         dHeadFireONDelay_cmm_H7 : DInt;   // Head#x fire ON delay [mm/100] {mm/100|mm|-50|50|O} / Head #7 fire ON delay [mm/100] {mm/100|mm|-50|50|O}
         dHeadFireOFFDelay_cmm_H7 : DInt;   // Head#x fire OFF delay [mm/100] {mm/100|mm|-50|50|O} / Head #7 fire OFF delay [mm/100] {mm/100|mm|-50|50|O}
         dHeadPressure_mN_H7 : DInt;   // Head#x pressure value [N/1000] {N/1000|N|16|180|O} / Head #7 pressure value [N/1000] {N/1000|N|16|180|O}
         dHeadFireONReaction_ms_H8 : DInt;   // Head#x fire ON reaction time [ms] {ms|s|0|1|M} / Head #8 fire ON reaction time [ms] {ms|s|0|1|M}
         dHeadFireOFFReaction_ms_H8 : DInt;   // Head#x fire OFF reaction time [ms] {ms|s|0|1|M} / Head #8 fire OFF reaction time [ms] {ms|s|0|1|M}
         dHeadOilONDelay_ms_H8 : DInt;   // Head#x Oil ON delay [ms]{ms|s|-2|2|O} / Head #8 Oil ON delay [ms]{ms|s|-2|2|O}
         dHeadOilOFFDelay_ms_H8 : DInt;   // Head#x Oil OFF delay [ms]{ms|s|-2|2|O} / Head #8 Oil OFF delay [ms]{ms|s|-2|2|O}
         dHeadFireONDelay_cmm_H8 : DInt;   // Head#x fire ON delay [mm/100] {mm/100|mm|-50|50|O} / Head #8 fire ON delay [mm/100] {mm/100|mm|-50|50|O}
         dHeadFireOFFDelay_cmm_H8 : DInt;   // Head#x fire OFF delay [mm/100] {mm/100|mm|-50|50|O} / Head #8 fire OFF delay [mm/100] {mm/100|mm|-50|50|O}
         dHeadPressure_mN_H8 : DInt;   // Head#x pressure value [N/1000] {N/1000|N|16|180|O} / Head #8 pressure value [N/1000] {N/1000|N|16|180|O}
         dSpare56 : DInt;
         dSpare57 : DInt;
         dSpare58 : DInt;
         dSpare59 : DInt;
         rSpare0 : Real;
         rSpare1 : Real;
         rSpare2 : Real;
         rSpare3 : Real;
         rSpare4 : Real;
         rSpare5 : Real;
         rSpare6 : Real;
         rSpare7 : Real;
         rSpare8 : Real;
         tManCmd : Struct
            xMan_FireON_H1 : Bool;   // Head#x manual fire ON {x|x|x|x|O} / Head #1 manual fire ON {x|x|x|x|O}
            xMan_FireOFF_H1 : Bool;   // Head#x manual fire OFF {x|x|x|x|O} / Head #1 manual fire OFF {x|x|x|x|O}
            xMan_OilON_H1 : Bool;   // Head#x manual oil ON {x|x|x|x|O} / Head #1 manual oil ON {x|x|x|x|O}
            xMan_FireON_H2 : Bool;   // Head#x manual fire ON {x|x|x|x|O} / Head #2 manual fire ON {x|x|x|x|O}
            xMan_FireOFF_H2 : Bool;   // Head#x manual fire OFF {x|x|x|x|O} / Head #2 manual fire OFF {x|x|x|x|O}
            xMan_OilON_H2 : Bool;   // Head#x manual oil ON {x|x|x|x|O} / Head #2 manual oil ON {x|x|x|x|O}
            xMan_FireON_H3 : Bool;   // Head#x manual fire ON {x|x|x|x|O} / Head #3 manual fire ON {x|x|x|x|O}
            xMan_FireOFF_H3 : Bool;   // Head#x manual fire OFF {x|x|x|x|O} / Head #3 manual fire OFF {x|x|x|x|O}
            xMan_OilON_H3 : Bool;   // Head#x manual oil ON {x|x|x|x|O} / Head #3 manual oil ON {x|x|x|x|O}
            xMan_FireON_H4 : Bool;   // Head#x manual fire ON {x|x|x|x|O} / Head #4 manual fire ON {x|x|x|x|O}
            xMan_FireOFF_H4 : Bool;   // Head#x manual fire OFF {x|x|x|x|O} / Head #4 manual fire OFF {x|x|x|x|O}
            xMan_OilON_H4 : Bool;   // Head#x manual oil ON {x|x|x|x|O} / Head #4 manual oil ON {x|x|x|x|O}
            xMan_FireON_H5 : Bool;   // Head#x manual fire ON {x|x|x|x|O} / Head #5 manual fire ON {x|x|x|x|O}
            xMan_FireOFF_H5 : Bool;   // Head#x manual fire OFF {x|x|x|x|O} / Head #5 manual fire OFF {x|x|x|x|O}
            xMan_OilON_H5 : Bool;   // Head#x manual oil ON {x|x|x|x|O} / Head #5 manual oil ON {x|x|x|x|O}
            xMan_FireON_H6 : Bool;   // Head#x manual fire ON {x|x|x|x|O} / Head #6 manual fire ON {x|x|x|x|O}
            xMan_FireOFF_H6 : Bool;   // Head#x manual fire OFF {x|x|x|x|O} / Head #6 manual fire OFF {x|x|x|x|O}
            xMan_OilON_H6 : Bool;   // Head#x manual oil ON {x|x|x|x|O} / Head #6 manual oil ON {x|x|x|x|O}
            xMan_FireON_H7 : Bool;   // Head#x manual fire ON {x|x|x|x|O} / Head #7 manual fire ON {x|x|x|x|O}
            xMan_FireOFF_H7 : Bool;   // Head#x manual fire OFF {x|x|x|x|O} / Head #7 manual fire OFF {x|x|x|x|O}
            xMan_OilON_H7 : Bool;   // Head#x manual oil ON {x|x|x|x|O} / Head #7 manual oil ON {x|x|x|x|O}
            xMan_FireON_H8 : Bool;   // Head#x manual fire ON {x|x|x|x|O} / Head #8 manual fire ON {x|x|x|x|O}
            xMan_FireOFF_H8 : Bool;   // Head#x manual fire OFF {x|x|x|x|O} / Head #8 manual fire OFF {x|x|x|x|O}
            xMan_OilON_H8 : Bool;   // Head#x manual oil ON {x|x|x|x|O} / Head #8 manual oil ON {x|x|x|x|O}
            xSpare24 : Bool;
            xSpare25 : Bool;
            xSpare26 : Bool;
            xSpare27 : Bool;
            xSpare28 : Bool;
            xSpare29 : Bool;
            xSpare30 : Bool;
            xSpare31 : Bool;
         END_STRUCT;
      END_STRUCT;
   END_VAR
BEGIN
END_DATA_BLOCK

DATA_BLOCK "DB_M256A_Scada"   // DB2013
{ S7_Optimized_Access := 'FALSE' }
VERSION : 0.1
   VAR
      tAlm : Struct   // HMI Alarms
         tE : Struct
            x0 : Bool;   // KE.Main emergency on
            x1 : Bool;   // KE1.Local emergency on
            x2 : Bool;   // Cabinet.Emergency localization
            x3 : Bool;   // SB1.Emergency localization
            x4 : Bool;   // SB2.Emergency localization
            x5 : Bool;
            x6 : Bool;
            x7 : Bool;
            x8 : Bool;
            x9 : Bool;
            x10 : Bool;
            x11 : Bool;
            x12 : Bool;
            x13 : Bool;
            x14 : Bool;
            x15 : Bool;
            x16 : Bool;
            x17 : Bool;
            x18 : Bool;
            x19 : Bool;
            x20 : Bool;
            x21 : Bool;
            x22 : Bool;
            x23 : Bool;
            x24 : Bool;
            x25 : Bool;
            x26 : Bool;
            x27 : Bool;
            x28 : Bool;
            x29 : Bool;
            x30 : Bool;
            x31 : Bool;
         END_STRUCT;
         tS : Struct
            tS0 : Struct
               x0 : Bool;   // Head#x carriage not in working position / Head#1 carriage not in working position
               x1 : Bool;   // Head#x carriage not in working position
               x2 : Bool;   // Head#x carriage not in working position
               x3 : Bool;   // Head#x carriage not in working position
               x4 : Bool;   // Head#x carriage not in working position
               x5 : Bool;   // Head#x carriage not in working position
               x6 : Bool;   // Head#x carriage not in working position
               x7 : Bool;   // Head#x carriage not in working position
               x8 : Bool;   // xB21QF1.Power supply 24V logic
               x9 : Bool;   // Head#x carriage not in working position / Head#2carriage not in working position
               x10 : Bool;   // Syncro.Main line meter gap outside the limits
               x11 : Bool;
               x12 : Bool;
               x13 : Bool;
               x14 : Bool;
               x15 : Bool;
               x16 : Bool;
               x17 : Bool;
               x18 : Bool;   // Head#x carriage not in working position / Head#3carriage not in working position
               x19 : Bool;
               x20 : Bool;
               x21 : Bool;
               x22 : Bool;
               x23 : Bool;
               x24 : Bool;
               x25 : Bool;
               x26 : Bool;
               x27 : Bool;
               x28 : Bool;
               x29 : Bool;
               x30 : Bool;
               x31 : Bool;
            END_STRUCT;
            tS1 : Struct
               x0 : Bool;   // Head#x carriage not in working position / Head#4carriage not in working position
               x1 : Bool;   // Syncro.YCut meter gap outside the limits
               x2 : Bool;
               x3 : Bool;
               x4 : Bool;
               x5 : Bool;
               x6 : Bool;
               x7 : Bool;
               x8 : Bool;   // xB21QF1.Power supply 24V logic
               x9 : Bool;   // Head#x carriage not in working position / Head#5carriage not in working position
               x10 : Bool;   // Syncro.Main line meter gap outside the limits
               x11 : Bool;
               x12 : Bool;
               x13 : Bool;
               x14 : Bool;
               x15 : Bool;
               x16 : Bool;
               x17 : Bool;
               x18 : Bool;   // Head#x carriage not in working position / Head#6carriage not in working position
               x19 : Bool;
               x20 : Bool;
               x21 : Bool;
               x22 : Bool;
               x23 : Bool;
               x24 : Bool;
               x25 : Bool;
               x26 : Bool;
               x27 : Bool;
               x28 : Bool;
               x29 : Bool;
               x30 : Bool;
               x31 : Bool;
            END_STRUCT;
            tS2 : Struct
               x0 : Bool;   // Head#x carriage not in working position / Head#7carriage not in working position
               x1 : Bool;   // Syncro.YCut meter gap outside the limits
               x2 : Bool;
               x3 : Bool;
               x4 : Bool;
               x5 : Bool;
               x6 : Bool;
               x7 : Bool;
               x8 : Bool;   // xB21QF1.Power supply 24V logic
               x9 : Bool;   // Head#x carriage not in working position / Head#8carriage not in working position
               x10 : Bool;   // Syncro.Main line meter gap outside the limits
               x11 : Bool;
               x12 : Bool;
               x13 : Bool;
               x14 : Bool;
               x15 : Bool;
               x16 : Bool;
               x17 : Bool;
               x18 : Bool;
               x19 : Bool;
               x20 : Bool;
               x21 : Bool;
               x22 : Bool;
               x23 : Bool;
               x24 : Bool;
               x25 : Bool;
               x26 : Bool;
               x27 : Bool;
               x28 : Bool;
               x29 : Bool;
               x30 : Bool;
               x31 : Bool;
            END_STRUCT;
            tS3 : Struct
               x0 : Bool;
               x1 : Bool;   // Syncro.YCut meter gap outside the limits
               x2 : Bool;
               x3 : Bool;
               x4 : Bool;
               x5 : Bool;
               x6 : Bool;
               x7 : Bool;
               x8 : Bool;   // xB21QF1.Power supply 24V logic
               x9 : Bool;
               x10 : Bool;   // Syncro.Main line meter gap outside the limits
               x11 : Bool;
               x12 : Bool;
               x13 : Bool;
               x14 : Bool;
               x15 : Bool;
               x16 : Bool;
               x17 : Bool;
               x18 : Bool;
               x19 : Bool;
               x20 : Bool;
               x21 : Bool;
               x22 : Bool;
               x23 : Bool;
               x24 : Bool;
               x25 : Bool;
               x26 : Bool;
               x27 : Bool;
               x28 : Bool;
               x29 : Bool;
               x30 : Bool;
               x31 : Bool;
            END_STRUCT;
         END_STRUCT;
         tF : Struct
            x0 : Bool;
            x1 : Bool;
            x2 : Bool;
            x3 : Bool;
            x4 : Bool;
            x5 : Bool;
            x6 : Bool;
            x7 : Bool;
            x8 : Bool;
            x9 : Bool;
            x10 : Bool;
            x11 : Bool;
            x12 : Bool;
            x13 : Bool;
            x14 : Bool;
            x15 : Bool;
            x16 : Bool;
            x17 : Bool;
            x18 : Bool;
            x19 : Bool;
            x20 : Bool;
            x21 : Bool;
            x22 : Bool;
            x23 : Bool;
            x24 : Bool;
            x25 : Bool;
            x26 : Bool;
            x27 : Bool;
            x28 : Bool;
            x29 : Bool;
            x30 : Bool;
            x31 : Bool;
         END_STRUCT;
         tW : Struct
            x0 : Bool;   // PLCA.Timeout receiving consumed message
            x1 : Bool;   // PLCB.Timeout receiving consumed message
            x2 : Bool;   // PLCA.Mission packet lost
            x3 : Bool;   // PLCB.Mission packet lost
            x4 : Bool;   // PLCA.Syncro packet lost
            x5 : Bool;   // PLCB.Syncro packet lost
            x6 : Bool;   // QF.Protection air conditioners
            x7 : Bool;
            x8 : Bool;
            x9 : Bool;
            x10 : Bool;
            x11 : Bool;
            x12 : Bool;
            x13 : Bool;
            x14 : Bool;
            x15 : Bool;
            x16 : Bool;
            x17 : Bool;
            x18 : Bool;
            x19 : Bool;
            x20 : Bool;
            x21 : Bool;
            x22 : Bool;
            x23 : Bool;
            x24 : Bool;
            x25 : Bool;
            x26 : Bool;
            x27 : Bool;
            x28 : Bool;
            x29 : Bool;
            x30 : Bool;
            x31 : Bool;
         END_STRUCT;
      END_STRUCT;
      tHMR : Struct   // HMI Read
         xSpare0 : Bool := FALSE;   // Calibration function allowed {x|x|x|x|O}
         xSpare1 : Bool;
         xSpare2 : Bool;
         xSpare3 : Bool;
         xSpare4 : Bool;
         xSpare5 : Bool;
         xSpare6 : Bool;
         xSpare7 : Bool;
         xSpare8 : Bool;
         xSpare9 : Bool;
         xSpare10 : Bool;
         xSpare11 : Bool;
         xSpare12 : Bool;
         xSpare13 : Bool;
         xSpare14 : Bool;
         xSpare15 : Bool := FALSE;
         xSpare16 : Bool;
         xSpare17 : Bool;
         xSpare18 : Bool;
         xSpare19 : Bool;
         xSpare20 : Bool;
         xSpare21 : Bool;
         xSpare22 : Bool;
         xSpare23 : Bool;
         xSpare24 : Bool;
         xSpare25 : Bool;
         xSpare26 : Bool;
         xSpare27 : Bool;
         xSpare28 : Bool;
         xSpare29 : Bool;
         xSpare30 : Bool;
         xSpare31 : Bool;
         xSpare : Array[0..15] of Bool;
         iSpare0 : Int;
         iSpare1 : Int;
         iSpare2 : Int;
         iSpare3 : Int;
         iSpare4 : Int;
         iSpare5 : Int;
         iSpare6 : Int;
         iSpare7 : Int;
         iSpare8 : Int;
         iSpare9 : Int;
         iSpare10 : Int;
         iSpare11 : Int;
         iSpare12 : Int;
         iSpare13 : Int;
         iSpare14 : Int;
         iSpare15 : Int;
         iSpare16 : Int;
         dHeadStatus_H1 : DInt;   // Head#x arming status (1=Up 3=Down 7=Anomaly) {x|x|x|x|O} / Head#1 arming status (1=Up 3=Down 7=Anomaly) {x|x|x|x|O}
         dHeadStatus_H2 : DInt;   // Head#x arming status (1=Up 3=Down 7=Anomaly) {x|x|x|x|O} / Head#2 arming status (1=Up 3=Down 7=Anomaly) {x|x|x|x|O}
         dHeadStatus_H3 : DInt;   // Head#x arming status (1=Up 3=Down 7=Anomaly) {x|x|x|x|O} / Head#3 arming status (1=Up 3=Down 7=Anomaly) {x|x|x|x|O}
         dHeadStatus_H4 : DInt;   // Head#x arming status (1=Up 3=Down 7=Anomaly) {x|x|x|x|O} / Head#4 arming status (1=Up 3=Down 7=Anomaly) {x|x|x|x|O}
         dHeadStatus_H5 : DInt;   // Head#x arming status (1=Up 3=Down 7=Anomaly) {x|x|x|x|O} / Head#5 arming status (1=Up 3=Down 7=Anomaly) {x|x|x|x|O}
         dHeadStatus_H6 : DInt;   // Head#x arming status (1=Up 3=Down 7=Anomaly) {x|x|x|x|O} / Head#6 arming status (1=Up 3=Down 7=Anomaly) {x|x|x|x|O}
         dHeadStatus_H7 : DInt;   // Head#x arming status (1=Up 3=Down 7=Anomaly) {x|x|x|x|O} / Head#7 arming status (1=Up 3=Down 7=Anomaly) {x|x|x|x|O}
         dHeadStatus_H8 : DInt;   // Head#x arming status (1=Up 3=Down 7=Anomaly) {x|x|x|x|O} / Head#8 arming status (1=Up 3=Down 7=Anomaly) {x|x|x|x|O}
         dSpare8 : DInt := 0;
         dSpare9 : DInt := 0;
         dSpare10 : DInt := 0;
         dSpare11 : DInt := 0;
         dSpare12 : DInt;
         dSpare13 : DInt;
         dSpare14 : DInt;
         dSpare15 : DInt;
         dSpare : Array[0..15] of DInt;
         rSpare0 : Real;
         rSpare1 : Real;
         rSpare2 : Real;
         rSpare3 : Real;
         rSpare4 : Real;
         rSpare5 : Real;
         rSpare6 : Real;
         rSpare7 : Real;
         rSpare8 : Real;
         tManCmd : Struct
            xMan_DescentFdbk_H1 : Bool;   // Head #x manual descent feedback {x|x|x|x|O} / Head #1 manual descent feedback {x|x|x|x|O}
            xMan_RiseFdbk_H1 : Bool;   // Head #x manual rise feedback {x|x|x|x|O} / Head #1 manual rise feedback {x|x|x|x|O}
            xMan_DescentFdbk_H2 : Bool;   // Head #x manual descent feedback {x|x|x|x|O} / Head #2 manual descent feedback {x|x|x|x|O}
            xMan_RiseFdbk_H2 : Bool;   // Head #x manual rise feedback {x|x|x|x|O} / Head #2 manual rise feedback {x|x|x|x|O}
            xMan_DescentFdbk_H3 : Bool;   // Head #x manual descent feedback {x|x|x|x|O} / Head #3 manual descent feedback {x|x|x|x|O}
            xMan_RiseFdbk_H3 : Bool;   // Head #x manual rise feedback {x|x|x|x|O} / Head #3 manual rise feedback {x|x|x|x|O}
            xMan_DescentFdbk_H4 : Bool;   // Head #x manual descent feedback {x|x|x|x|O} / Head #4 manual descent feedback {x|x|x|x|O}
            xMan_RiseFdbk_H4 : Bool;   // Head #x manual rise feedback {x|x|x|x|O} / Head #4 manual rise feedback {x|x|x|x|O}
            xMan_DescentFdbk_H5 : Bool;   // Head #x manual descent feedback {x|x|x|x|O} / Head #5 manual descent feedback {x|x|x|x|O}
            xMan_RiseFdbk_H5 : Bool;   // Head #x manual rise feedback {x|x|x|x|O} / Head #5 manual rise feedback {x|x|x|x|O}
            xMan_DescentFdbk_H6 : Bool;   // Head #x manual descent feedback {x|x|x|x|O} / Head #6 manual descent feedback {x|x|x|x|O}
            xMan_RiseFdbk_H6 : Bool;   // Head #x manual rise feedback {x|x|x|x|O} / Head #6 manual rise feedback {x|x|x|x|O}
            xMan_DescentFdbk_H7 : Bool;   // Head #x manual descent feedback {x|x|x|x|O} / Head #7 manual descent feedback {x|x|x|x|O}
            xMan_RiseFdbk_H7 : Bool;   // Head #x manual rise feedback {x|x|x|x|O} / Head #7 manual rise feedback {x|x|x|x|O}
            xMan_DescentFdbk_H8 : Bool;   // Head #x manual descent feedback {x|x|x|x|O} / Head #8 manual descent feedback {x|x|x|x|O}
            xMan_RiseFdbk_H8 : Bool;   // Head #x manual rise feedback {x|x|x|x|O} / Head #8 manual rise feedback {x|x|x|x|O}
            xSpare : Array[0..15] of Bool;
         END_STRUCT;
      END_STRUCT;
      tHMW : Struct   // HMI Write
         xSpare0 : Bool := FALSE;   // Automatic mode request {x|x|x|x|O}
         xSpare1 : Bool := FALSE;   // Manual mode request {x|x|x|x|O}
         xSpare2 : Bool := FALSE;   // Bridge out of production request {x|x|x|x|O}
         xSpare3 : Bool := FALSE;   // Bridge in production request {x|x|x|x|O}
         xSpare4 : Bool := FALSE;   // Cut during glass break {x|x|x|x|O}
         xSpare5 : Bool := FALSE;   // Motors and cards initialize {x|x|x|x|M}
         xSpare6 : Bool := FALSE;   // Force the homing of the heads {x|x|x|x|M}
         xSpare7 : Bool := FALSE;   // Position calibration request {x|x|x|x|M}
         xSpare8 : Bool := FALSE;   // Bridge offset calibration request {x|x|x|x|M}
         xSpare9 : Bool;
         xSpare10 : Bool;
         xSpare11 : Bool;
         xSpare12 : Bool;
         xSpare13 : Bool;
         xSpare14 : Bool := FALSE;
         xSpare15 : Bool := FALSE;
         xSpare16 : Bool := TRUE;
         xSpare17 : Bool := TRUE;
         xSpare18 : Bool := TRUE;
         xSpare19 : Bool := TRUE;
         xSpare20 : Bool := TRUE;
         xSpare21 : Bool := TRUE;
         xSpare22 : Bool := TRUE;
         xSpare23 : Bool := TRUE;
         xSpare24 : Bool;
         xSpare25 : Bool;
         xSpare26 : Bool;
         xSpare27 : Bool;
         xSpare28 : Bool;
         xSpare29 : Bool;
         xSpare30 : Bool;
         xSpare31 : Bool;
         xSpare : Array[0..15] of Bool;
         iSpare0 : Int;
         iSpare1 : Int;
         iSpare2 : Int;
         iSpare3 : Int;
         iSpare4 : Int;
         iSpare5 : Int;
         iSpare6 : Int;
         iSpare7 : Int;
         iSpare8 : Int;
         iSpare9 : Int;
         iSpare10 : Int;
         iSpare11 : Int;
         iSpare12 : Int;
         iSpare13 : Int;
         iSpare14 : Int;
         iSpare15 : Int;
         iSpare16 : Int := 0;
         dRaiseReactTime_ms_H1 : DInt;   // Head#x raise reaction time [ms] {ms|s|-200|200|M} / Head#1 raise reaction time [ms] {ms|s|-200|200|M}
         dDescentReactTime_ms_H1 : DInt;   // Head#x descent reaction time [ms] {ms|s|0|3000|M} / Head#1 descent reaction time [ms] {ms|s|0|3000|M}
         dRaiseReactTime_ms_H2 : DInt;   // Head#x raise reaction time [ms] {ms|s|-200|200|M} / Head#2 raise reaction time [ms] {ms|s|-200|200|M}
         dDescentReactTime_ms_H2 : DInt;   // Head#x descent reaction time [ms] {ms|s|0|3000|M} / Head#2 descent reaction time [ms] {ms|s|0|3000|M}
         dRaiseReactTime_ms_H3 : DInt;   // Head#x raise reaction time [ms] {ms|s|-200|200|M} / Head#3 raise reaction time [ms] {ms|s|-200|200|M}
         dDescentReactTime_ms_H3 : DInt;   // Head#x descent reaction time [ms] {ms|s|0|3000|M} / Head#3 descent reaction time [ms] {ms|s|0|3000|M}
         dRaiseReactTime_ms_H4 : DInt;   // Head#x raise reaction time [ms] {ms|s|-200|200|M} / Head#4 raise reaction time [ms] {ms|s|-200|200|M}
         dDescentReactTime_ms_H4 : DInt;   // Head#x descent reaction time [ms] {ms|s|0|3000|M} / Head#4 descent reaction time [ms] {ms|s|0|3000|M}
         dRaiseReactTime_ms_H5 : DInt;   // Head#x raise reaction time [ms] {ms|s|-200|200|M} / Head#5raise reaction time [ms] {ms|s|-200|200|M}
         dDescentReactTime_ms_H5 : DInt;   // Head#x descent reaction time [ms] {ms|s|0|3000|M} / Head#5descent reaction time [ms] {ms|s|0|3000|M}
         dRaiseReactTime_ms_H6 : DInt;   // Head#x raise reaction time [ms] {ms|s|-200|200|M} / Head#6 raise reaction time [ms] {ms|s|-200|200|M}
         dDescentReactTime_ms_H6 : DInt;   // Head#x descent reaction time [ms] {ms|s|0|3000|M} / Head#6 descent reaction time [ms] {ms|s|0|3000|M}
         dRaiseReactTime_ms_H7 : DInt;   // Head#x raise reaction time [ms] {ms|s|-200|200|M} / Head#7 raise reaction time [ms] {ms|s|-200|200|M}
         dDescentReactTime_ms_H7 : DInt;   // Head#x descent reaction time [ms] {ms|s|0|3000|M} / Head#7 descent reaction time [ms] {ms|s|0|3000|M}
         dRaiseReactTime_ms_H8 : DInt;   // Head#x raise reaction time [ms] {ms|s|-200|200|M} / Head#8 raise reaction time [ms] {ms|s|-200|200|M}
         dDescentReactTime_ms_H8 : DInt;   // Head#x descent reaction time [ms] {ms|s|0|3000|M} / Head#8 descent reaction time [ms] {ms|s|0|3000|M}
         dSpare16 : DInt;
         dSpare17 : DInt;
         dSpare18 : DInt;
         dSpare19 : DInt;
         dSpare20 : DInt;
         dSpare21 : DInt;
         dSpare22 : DInt;
         dSpare23 : DInt;
         dSpare24 : DInt;
         dSpare25 : DInt;
         dSpare26 : DInt;
         dSpare27 : DInt;
         dSpare28 : DInt;
         dSpare29 : DInt;
         dSpare30 : DInt;
         dSpare31 : DInt;
         dSpare32 : DInt;
         dSpare33 : DInt;
         dSpare34 : DInt;
         dSpare35 : DInt;
         dSpare36 : DInt;
         dSpare37 : DInt;
         dSpare38 : DInt;
         dSpare39 : DInt;
         dSpare : Array[0..19] of DInt;
         rSpare0 : Real;
         rSpare1 : Real;
         rSpare2 : Real;
         rSpare3 : Real;
         rSpare4 : Real;
         rSpare5 : Real;
         rSpare6 : Real;
         rSpare7 : Real;
         rSpare8 : Real;
         tManCmd : Struct
            xManDescent_H1 : Bool;   // Head #x manual Descent {x|x|x|x|O} / Head #1 manual Descent {x|x|x|x|O}
            xManRise_H1 : Bool;   // Head #x manual rise {x|x|x|x|O} / Head #1 manual rise {x|x|x|x|O}
            xManRise_H2 : Bool;   // Head #x manual rise {x|x|x|x|O} / Head #2 manual rise {x|x|x|x|O}
            xManDescent_H2 : Bool;   // Head #x manual Descent {x|x|x|x|O} / Head #2 manual Descent {x|x|x|x|O}
            xManRise_H3 : Bool;   // Head #x manual rise {x|x|x|x|O} / Head #3 manual rise {x|x|x|x|O}
            xManDescent_H3 : Bool;   // Head #x manual Descent {x|x|x|x|O} / Head #3 manual Descent {x|x|x|x|O}
            xManRise_H4 : Bool;   // Head #x manual rise {x|x|x|x|O} / Head #4 manual rise {x|x|x|x|O}
            xManDescent_H4 : Bool;   // Head #x manual Descent {x|x|x|x|O} / Head #4 manual Descent {x|x|x|x|O}
            xManRise_H5 : Bool;   // Head #x manual rise {x|x|x|x|O} / Head #5 manual rise {x|x|x|x|O}
            xManDescent_H5 : Bool;   // Head #x manual Descent {x|x|x|x|O} / Head #5 manual Descent {x|x|x|x|O}
            xManRise_H6 : Bool;   // Head #x manual rise {x|x|x|x|O} / Head #6 manual rise {x|x|x|x|O}
            xManDescent_H6 : Bool;   // Head #x manual Descent {x|x|x|x|O} / Head #6 manual Descent {x|x|x|x|O}
            xManRise_H7 : Bool;   // Head #x manual rise {x|x|x|x|O} / Head #7 manual rise {x|x|x|x|O}
            xManDescent_H7 : Bool;   // Head #x manual Descent {x|x|x|x|O} / Head #7 manual Descent {x|x|x|x|O}
            xManRise_H8 : Bool;   // Head #x manual rise {x|x|x|x|O} / Head #8 manual rise {x|x|x|x|O}
            xManDescent_H8 : Bool;   // Head #x manual Descent {x|x|x|x|O} / Head #8 manual Descent {x|x|x|x|O}
            xSpare16 : Bool;
            xSpare17 : Bool;
            xSpare18 : Bool;
            xSpare19 : Bool;
            xSpare20 : Bool;
            xSpare21 : Bool;
            xSpare22 : Bool;
            xSpare23 : Bool;
            xSpare24 : Bool;
            xSpare25 : Bool;
            xSpare26 : Bool;
            xSpare27 : Bool;
            xSpare28 : Bool;
            xSpare29 : Bool;
            xSpare30 : Bool;
            xSpare31 : Bool;
         END_STRUCT;
      END_STRUCT;
   END_VAR
BEGIN
END_DATA_BLOCK

DATA_BLOCK "DB_Scada_default"   // DB2112
{ S7_Optimized_Access := 'FALSE' }
VERSION : 0.1
   VAR
      tAlm : Struct   // HMI Alarms
         tE : Struct
            x0 : Bool;   // KE.Main emergency on
            x1 : Bool;   // KE1.Local emergency on
            x2 : Bool;   // Cabinet.Emergency localization
            x3 : Bool;   // SB1.Emergency localization
            x4 : Bool;   // SB2.Emergency localization
            x5 : Bool;
            x6 : Bool;
            x7 : Bool;
            x8 : Bool;
            x9 : Bool;
            x10 : Bool;
            x11 : Bool;
            x12 : Bool;
            x13 : Bool;
            x14 : Bool;
            x15 : Bool;
            x16 : Bool;
            x17 : Bool;
            x18 : Bool;
            x19 : Bool;
            x20 : Bool;
            x21 : Bool;
            x22 : Bool;
            x23 : Bool;
            x24 : Bool;
            x25 : Bool;
            x26 : Bool;
            x27 : Bool;
            x28 : Bool;
            x29 : Bool;
            x30 : Bool;
            x31 : Bool;
         END_STRUCT;
         tS : Struct
            tS0 : Struct
               x0 : Bool;
               x1 : Bool;   // Syncro.YCut meter gap outside the limits
               x2 : Bool;
               x3 : Bool;
               x4 : Bool;
               x5 : Bool;
               x6 : Bool;
               x7 : Bool;
               x8 : Bool;   // xB21QF1.Power supply 24V logic
               x9 : Bool;
               x10 : Bool;   // Syncro.Main line meter gap outside the limits
               x11 : Bool;
               x12 : Bool;
               x13 : Bool;
               x14 : Bool;
               x15 : Bool;
               x16 : Bool;
               x17 : Bool;
               x18 : Bool;
               x19 : Bool;
               x20 : Bool;
               x21 : Bool;
               x22 : Bool;
               x23 : Bool;
               x24 : Bool;
               x25 : Bool;
               x26 : Bool;
               x27 : Bool;
               x28 : Bool;
               x29 : Bool;
               x30 : Bool;
               x31 : Bool;
            END_STRUCT;
            tS1 : Struct
               x0 : Bool;
               x1 : Bool;   // Syncro.YCut meter gap outside the limits
               x2 : Bool;
               x3 : Bool;
               x4 : Bool;
               x5 : Bool;
               x6 : Bool;
               x7 : Bool;
               x8 : Bool;   // xB21QF1.Power supply 24V logic
               x9 : Bool;
               x10 : Bool;   // Syncro.Main line meter gap outside the limits
               x11 : Bool;
               x12 : Bool;
               x13 : Bool;
               x14 : Bool;
               x15 : Bool;
               x16 : Bool;
               x17 : Bool;
               x18 : Bool;
               x19 : Bool;
               x20 : Bool;
               x21 : Bool;
               x22 : Bool;
               x23 : Bool;
               x24 : Bool;
               x25 : Bool;
               x26 : Bool;
               x27 : Bool;
               x28 : Bool;
               x29 : Bool;
               x30 : Bool;
               x31 : Bool;
            END_STRUCT;
            tS2 : Struct
               x0 : Bool;
               x1 : Bool;   // Syncro.YCut meter gap outside the limits
               x2 : Bool;
               x3 : Bool;
               x4 : Bool;
               x5 : Bool;
               x6 : Bool;
               x7 : Bool;
               x8 : Bool;   // xB21QF1.Power supply 24V logic
               x9 : Bool;
               x10 : Bool;   // Syncro.Main line meter gap outside the limits
               x11 : Bool;
               x12 : Bool;
               x13 : Bool;
               x14 : Bool;
               x15 : Bool;
               x16 : Bool;
               x17 : Bool;
               x18 : Bool;
               x19 : Bool;
               x20 : Bool;
               x21 : Bool;
               x22 : Bool;
               x23 : Bool;
               x24 : Bool;
               x25 : Bool;
               x26 : Bool;
               x27 : Bool;
               x28 : Bool;
               x29 : Bool;
               x30 : Bool;
               x31 : Bool;
            END_STRUCT;
            tS3 : Struct
               x0 : Bool;
               x1 : Bool;   // Syncro.YCut meter gap outside the limits
               x2 : Bool;
               x3 : Bool;
               x4 : Bool;
               x5 : Bool;
               x6 : Bool;
               x7 : Bool;
               x8 : Bool;   // xB21QF1.Power supply 24V logic
               x9 : Bool;
               x10 : Bool;   // Syncro.Main line meter gap outside the limits
               x11 : Bool;
               x12 : Bool;
               x13 : Bool;
               x14 : Bool;
               x15 : Bool;
               x16 : Bool;
               x17 : Bool;
               x18 : Bool;
               x19 : Bool;
               x20 : Bool;
               x21 : Bool;
               x22 : Bool;
               x23 : Bool;
               x24 : Bool;
               x25 : Bool;
               x26 : Bool;
               x27 : Bool;
               x28 : Bool;
               x29 : Bool;
               x30 : Bool;
               x31 : Bool;
            END_STRUCT;
         END_STRUCT;
         tF : Struct
            x0 : Bool;
            x1 : Bool;
            x2 : Bool;
            x3 : Bool;
            x4 : Bool;
            x5 : Bool;
            x6 : Bool;
            x7 : Bool;
            x8 : Bool;
            x9 : Bool;
            x10 : Bool;
            x11 : Bool;
            x12 : Bool;
            x13 : Bool;
            x14 : Bool;
            x15 : Bool;
            x16 : Bool;
            x17 : Bool;
            x18 : Bool;
            x19 : Bool;
            x20 : Bool;
            x21 : Bool;
            x22 : Bool;
            x23 : Bool;
            x24 : Bool;
            x25 : Bool;
            x26 : Bool;
            x27 : Bool;
            x28 : Bool;
            x29 : Bool;
            x30 : Bool;
            x31 : Bool;
         END_STRUCT;
         tW : Struct
            x0 : Bool;   // PLCA.Timeout receiving consumed message
            x1 : Bool;   // PLCB.Timeout receiving consumed message
            x2 : Bool;   // PLCA.Mission packet lost
            x3 : Bool;   // PLCB.Mission packet lost
            x4 : Bool;   // PLCA.Syncro packet lost
            x5 : Bool;   // PLCB.Syncro packet lost
            x6 : Bool;   // QF.Protection air conditioners
            x7 : Bool;
            x8 : Bool;
            x9 : Bool;
            x10 : Bool;
            x11 : Bool;
            x12 : Bool;
            x13 : Bool;
            x14 : Bool;
            x15 : Bool;
            x16 : Bool;
            x17 : Bool;
            x18 : Bool;
            x19 : Bool;
            x20 : Bool;
            x21 : Bool;
            x22 : Bool;
            x23 : Bool;
            x24 : Bool;
            x25 : Bool;
            x26 : Bool;
            x27 : Bool;
            x28 : Bool;
            x29 : Bool;
            x30 : Bool;
            x31 : Bool;
         END_STRUCT;
      END_STRUCT;
      tHMR : Struct   // HMI Read
         xSpare0 : Bool := FALSE;   // Calibration function allowed {x|x|x|x|O}
         xSpare1 : Bool;
         xSpare2 : Bool;
         xSpare3 : Bool;
         xSpare4 : Bool;
         xSpare5 : Bool;
         xSpare6 : Bool;
         xSpare7 : Bool;
         xSpare8 : Bool;
         xSpare9 : Bool;
         xSpare10 : Bool;
         xSpare11 : Bool;
         xSpare12 : Bool;
         xSpare13 : Bool;
         xSpare14 : Bool;
         xSpare15 : Bool := FALSE;
         xSpare16 : Bool;
         xSpare17 : Bool;
         xSpare18 : Bool;
         xSpare19 : Bool;
         xSpare20 : Bool;
         xSpare21 : Bool;
         xSpare22 : Bool;
         xSpare23 : Bool;
         xSpare24 : Bool;
         xSpare25 : Bool;
         xSpare26 : Bool;
         xSpare27 : Bool;
         xSpare28 : Bool;
         xSpare29 : Bool;
         xSpare30 : Bool;
         xSpare31 : Bool;
         xSpare : Array[0..15] of Bool;
         iSpare0 : Int;
         iSpare1 : Int;
         iSpare2 : Int;
         iSpare3 : Int;
         iSpare4 : Int;
         iSpare5 : Int;
         iSpare6 : Int;
         iSpare7 : Int;
         iSpare8 : Int;
         iSpare9 : Int;
         iSpare10 : Int;
         iSpare11 : Int;
         iSpare12 : Int;
         iSpare13 : Int;
         iSpare14 : Int;
         iSpare15 : Int;
         iSpare16 : Int;
         dSpare0 : DInt := 0;   // Zone modality (1=Manual;4=Automatic;8=Manual request) {x|x|x|x|O}
         dSpare1 : DInt := 0;   // HMI Alarms
         dSpare2 : DInt := 0;   // HMI Write
         dSpare3 : DInt := 0;   // Production modality request (1=Out of Production 3= In production) {x|x|x|x|O}
         dSpare4 : DInt := 0;   // Production modality actual (1=Out of production 3=In production 8=Out of production request 9=In production request) {x|x|x|x|O}
         dSpare5 : DInt := 0;
         dSpare6 : DInt := 0;
         dSpare7 : DInt := 0;
         dSpare8 : DInt := 0;
         dSpare9 : DInt := 0;
         dSpare10 : DInt := 0;
         dSpare11 : DInt := 0;
         dSpare12 : DInt;
         dSpare13 : DInt;
         dSpare14 : DInt;
         dSpare15 : DInt;
         dSpare : Array[0..15] of DInt;
         rSpare0 : Real;
         rSpare1 : Real;
         rSpare2 : Real;
         rSpare3 : Real;
         rSpare4 : Real;
         rSpare5 : Real;
         rSpare6 : Real;
         rSpare7 : Real;
         rSpare8 : Real;
         tManCmd : Struct
            xSpare0 : Bool;
            xSpare1 : Bool;
            xSpare2 : Bool;
            xSpare3 : Bool;
            xSpare4 : Bool;
            xSpare5 : Bool;
            xSpare6 : Bool;
            xSpare7 : Bool;
            xSpare8 : Bool;
            xSpare9 : Bool;
            xSpare10 : Bool;
            xSpare11 : Bool;
            xSpare12 : Bool;
            xSpare13 : Bool;
            xSpare14 : Bool;
            xSpare15 : Bool;
            xSpare : Array[0..15] of Bool;
         END_STRUCT;
      END_STRUCT;
      tHMW : Struct   // HMI Write
         xSpare0 : Bool := FALSE;   // Automatic mode request {x|x|x|x|O}
         xSpare1 : Bool := FALSE;   // Manual mode request {x|x|x|x|O}
         xSpare2 : Bool := FALSE;   // Bridge out of production request {x|x|x|x|O}
         xSpare3 : Bool := FALSE;   // Bridge in production request {x|x|x|x|O}
         xSpare4 : Bool := FALSE;   // Cut during glass break {x|x|x|x|O}
         xSpare5 : Bool := FALSE;   // Motors and cards initialize {x|x|x|x|M}
         xSpare6 : Bool := FALSE;   // Force the homing of the heads {x|x|x|x|M}
         xSpare7 : Bool := FALSE;   // Position calibration request {x|x|x|x|M}
         xSpare8 : Bool := FALSE;   // Bridge offset calibration request {x|x|x|x|M}
         xSpare9 : Bool;
         xSpare10 : Bool;
         xSpare11 : Bool;
         xSpare12 : Bool;
         xSpare13 : Bool;
         xSpare14 : Bool := FALSE;
         xSpare15 : Bool := FALSE;
         xSpare16 : Bool := TRUE;
         xSpare17 : Bool := TRUE;
         xSpare18 : Bool := TRUE;
         xSpare19 : Bool := TRUE;
         xSpare20 : Bool := TRUE;
         xSpare21 : Bool := TRUE;
         xSpare22 : Bool := TRUE;
         xSpare23 : Bool := TRUE;
         xSpare24 : Bool;
         xSpare25 : Bool;
         xSpare26 : Bool;
         xSpare27 : Bool;
         xSpare28 : Bool;
         xSpare29 : Bool;
         xSpare30 : Bool;
         xSpare31 : Bool;
         xSpare : Array[0..15] of Bool;
         iSpare0 : Int;
         iSpare1 : Int;
         iSpare2 : Int;
         iSpare3 : Int;
         iSpare4 : Int;
         iSpare5 : Int;
         iSpare6 : Int;
         iSpare7 : Int;
         iSpare8 : Int;
         iSpare9 : Int;
         iSpare10 : Int;
         iSpare11 : Int;
         iSpare12 : Int;
         iSpare13 : Int;
         iSpare14 : Int;
         iSpare15 : Int;
         iSpare16 : Int := 0;
         dSpare0 : DInt := 0;   // Calibration. number of lite on calibration {x|x|1|8|M}
         dSpare1 : DInt := 0;   // Calibration. Move all the heads of this offset {mm/100|mm|-100|100|M}
         dSpare2 : DInt := 0;   // Pressure scaler during sample plate [%] {%|%|0|100|O}
         dSpare3 : DInt := 0;
         dSpare4 : DInt;
         dSpare5 : DInt;
         dSpare6 : DInt;
         dSpare7 : DInt;
         dSpare8 : DInt;
         dSpare9 : DInt;
         dSpare10 : DInt;
         dSpare11 : DInt;
         dSpare12 : DInt;
         dSpare13 : DInt;
         dSpare14 : DInt;
         dSpare15 : DInt;
         dSpare16 : DInt;
         dSpare17 : DInt;
         dSpare18 : DInt;
         dSpare19 : DInt;
         dSpare20 : DInt;
         dSpare21 : DInt;
         dSpare22 : DInt;
         dSpare23 : DInt;
         dSpare24 : DInt;
         dSpare25 : DInt;
         dSpare26 : DInt;
         dSpare27 : DInt;
         dSpare28 : DInt;
         dSpare29 : DInt;
         dSpare30 : DInt;
         dSpare31 : DInt;
         dSpare32 : DInt;
         dSpare33 : DInt;
         dSpare34 : DInt;
         dSpare35 : DInt;
         dSpare36 : DInt;
         dSpare37 : DInt;
         dSpare38 : DInt;
         dSpare39 : DInt;
         dSpare : Array[0..19] of DInt;
         rSpare0 : Real;
         rSpare1 : Real;
         rSpare2 : Real;
         rSpare3 : Real;
         rSpare4 : Real;
         rSpare5 : Real;
         rSpare6 : Real;
         rSpare7 : Real;
         rSpare8 : Real;
         tManCmd : Struct
            xSpare0 : Bool := FALSE;
            xSpare1 : Bool := FALSE;
            xSpare2 : Bool;
            xSpare3 : Bool;
            xSpare4 : Bool;
            xSpare5 : Bool;
            xSpare6 : Bool;
            xSpare7 : Bool;
            xSpare8 : Bool;
            xSpare9 : Bool;
            xSpare10 : Bool;
            xSpare11 : Bool;
            xSpare12 : Bool;
            xSpare13 : Bool;
            xSpare14 : Bool;
            xSpare15 : Bool;
            xSpare16 : Bool;
            xSpare17 : Bool;
            xSpare18 : Bool;
            xSpare19 : Bool;
            xSpare20 : Bool;
            xSpare21 : Bool;
            xSpare22 : Bool;
            xSpare23 : Bool;
            xSpare24 : Bool;
            xSpare25 : Bool;
            xSpare26 : Bool;
            xSpare27 : Bool;
            xSpare28 : Bool;
            xSpare29 : Bool;
            xSpare30 : Bool;
            xSpare31 : Bool;
         END_STRUCT;
      END_STRUCT;
   END_VAR
BEGIN
END_DATA_BLOCK

// folder: Communication

DATA_BLOCK "CM_Manager"   // DB1
{ S7_Optimized_Access := 'TRUE' }
VERSION : 0.1
BEGIN
END_DATA_BLOCK

DATA_BLOCK "CM_IDEV_FromMainLine"   // DB2
{ S7_Optimized_Access := 'TRUE' }
VERSION : 0.1
BEGIN
END_DATA_BLOCK

DATA_BLOCK "CM_IDEV_ToMainLine"   // DB3
{ S7_Optimized_Access := 'TRUE' }
VERSION : 0.1
BEGIN
END_DATA_BLOCK

DATA_BLOCK "CM_RECV_MissionData"   // DB4
{ S7_Optimized_Access := 'TRUE' }
VERSION : 0.1
BEGIN
END_DATA_BLOCK

DATA_BLOCK "CM_RECV_SyncroData"   // DB8
{ S7_Optimized_Access := 'TRUE' }
VERSION : 0.1
BEGIN
END_DATA_BLOCK

DATA_BLOCK "CM_BRCV_FromMainLine0"   // DB12
{ S7_Optimized_Access := 'TRUE' }
VERSION : 0.1
BEGIN
END_DATA_BLOCK

DATA_BLOCK "CM_BRCV_FromMainLine1"   // DB24
{ S7_Optimized_Access := 'TRUE' }
VERSION : 0.1
BEGIN
END_DATA_BLOCK

// folder: ILx2_Blocks

DATA_BLOCK "ILx2T_Parameter_Initialize_DB"   // DB10
{ S7_Optimized_Access := 'TRUE' }
VERSION : 1.1
// stored: InstanceOfName ILx2T_Parameter_Read_Write
"ILx2T_Parameter_Read_Write"
BEGIN
END_DATA_BLOCK

// folder: Subroutine

DATA_BLOCK "OB_Initialize"   // DB18
{ S7_Optimized_Access := 'TRUE' }
AUTHOR : Cigliutt
FAMILY : GP
VERSION : 1.0
// stored: InstanceOfName GP_OB_Initialize
"GP_OB_Initialize"
BEGIN
END_DATA_BLOCK

// folder: TaskErrors

DATA_BLOCK "RALRM_AUX_DB"   // DB59
{ S7_Optimized_Access := 'TRUE' }
VERSION : 0.1
   VAR RETAIN
      tAlm : Struct   // HMI Alarms
         tS : Struct   // Stopping faults
            xSpare_0 : Bool := FALSE;
            xSpare_1 : Bool := FALSE;
            xSpare_2 : Bool := FALSE;
            xSpare_3 : Bool := FALSE;
            xSpare_4 : Bool := FALSE;
            xSpare_5 : Bool := FALSE;
            xSpare_6 : Bool := FALSE;
            xSpare_7 : Bool := FALSE;
            xSpare_8 : Bool := FALSE;
            xSpare_9 : Bool := FALSE;
            xSpare_10 : Bool := FALSE;
            xSpare_11 : Bool := FALSE;
            xSpare_12 : Bool := FALSE;
            xSpare_13 : Bool := FALSE;
            xSpare_14 : Bool := FALSE;
            xSpare_15 : Bool := FALSE;
            xSpare_16 : Bool := FALSE;
            xSpare_17 : Bool := FALSE;
            xSpare_18 : Bool := FALSE;
            xSpare_19 : Bool := FALSE;
            xSpare_20 : Bool := FALSE;
            xSpare_21 : Bool := FALSE;
            xSpare_22 : Bool := FALSE;
            xSpare_23 : Bool := FALSE;
            xSpare_24 : Bool := FALSE;
            xSpare_25 : Bool := FALSE;
            xSpare_26 : Bool := FALSE;
            xSpare_27 : Bool := FALSE;
            xSpare_28 : Bool := FALSE;
            xSpare_29 : Bool := FALSE;
            xSpare_30 : Bool := FALSE;
            xSpare_31 : Bool := FALSE;
         END_STRUCT;
         tF : Struct   // Faults
            xDevice1 : Bool := FALSE;   // R13QF1.R13QF2.Power failure 230v auxiliary / Status device error.Device#1
            xDevice2 : Bool := FALSE;   // R18QF3.Power supply 24v logic / Status device error.Device#2
            xDevice3 : Bool := FALSE;   // R18QF4.Power supply 24v logic / Status device error.Device#3
            xDevice4 : Bool := FALSE;   // R18AP1.Redundancy 24v ok / Status device error.Device#4
            xDevice5 : Bool := FALSE;   // Status device error.Device#5
            xDevice6 : Bool := FALSE;   // Status device error.Device#6
            xDevice7 : Bool := FALSE;   // Status device error.Device#7
            xDevice8 : Bool := FALSE;   // Status device error.Device#8
            xDevice9 : Bool := FALSE;   // Status device error.Device#9
            xDevice10 : Bool := FALSE;   // Status device error.Device#10
            xSpare_10 : Bool := FALSE;
            xSpare_11 : Bool := FALSE;
            xSpare_12 : Bool;
            xSpare_13 : Bool;   // M250.R12KM1.Feedback rotation
            xSpare_14 : Bool;
            xSpare_15 : Bool;
            xSpare_16 : Bool;
            xSpare_17 : Bool;   // R204SP1.Compressed air presence cutting bridges
            xSpare_18 : Bool;
            xSpare_19 : Bool;
            xSpare_20 : Bool := FALSE;
            xSpare_21 : Bool := FALSE;
            xSpare_22 : Bool := FALSE;
            xSpare_23 : Bool := FALSE;
            xSpare_24 : Bool := FALSE;
            xSpare_25 : Bool := FALSE;
            xSpare_26 : Bool := FALSE;
            xSpare_27 : Bool := FALSE;
            xSpare_28 : Bool := FALSE;
            xSpare_29 : Bool := FALSE;
            xSpare_30 : Bool := FALSE;
            xSpare_31 : Bool := FALSE;
         END_STRUCT;
         tW : Struct   // Warnings
            xSpare_0 : Bool := FALSE;
            xSpare_1 : Bool := FALSE;
            xSpare_2 : Bool := FALSE;
            xSpare_3 : Bool := FALSE;
            xSpare_4 : Bool := FALSE;
            xSpare_5 : Bool := FALSE;
            xSpare_6 : Bool := FALSE;
            xSpare_7 : Bool := FALSE;
            xSpare_8 : Bool := FALSE;
            xSpare_9 : Bool := FALSE;
            xSpare_10 : Bool := FALSE;
            xSpare_11 : Bool := FALSE;
            xSpare_12 : Bool := FALSE;
            xSpare_13 : Bool := FALSE;
            xSpare_14 : Bool := FALSE;
            xSpare_15 : Bool := FALSE;
            xSpare_16 : Bool := FALSE;
            xSpare_17 : Bool := FALSE;
            xSpare_18 : Bool := FALSE;
            xSpare_19 : Bool := FALSE;
            xSpare_20 : Bool := FALSE;
            xSpare_21 : Bool := FALSE;
            xSpare_22 : Bool := FALSE;
            xSpare_23 : Bool := FALSE;
            xSpare_24 : Bool := FALSE;
            xSpare_25 : Bool := FALSE;
            xSpare_26 : Bool := FALSE;
            xSpare_27 : Bool := FALSE;
            xSpare_28 : Bool := FALSE;
            xSpare_29 : Bool := FALSE;
            xSpare_30 : Bool := FALSE;
            xSpare_31 : Bool := FALSE;
         END_STRUCT;
      END_STRUCT;
   END_VAR
BEGIN
END_DATA_BLOCK

// folder: (top level)

FUNCTION_BLOCK "M256_Manager"   // FB11, LAD
TITLE = #### HEAD MANAGER ####
{ S7_Optimized_Access := 'TRUE' }
VERSION : 0.1
   VAR_INPUT
      IN_tConnectionData : Array[0.."CONST_dNumberOfHeadsCycle"] of "UDT_MB_ConnData";   // IP and connection ID
   END_VAR
   VAR
      M256M_IDB : Array[0.."CONST_dNumberOfHeadsCycle"] of "M256M";
      M256F_IDB : Array[0.."CONST_dNumberOfHeadsCycle"] of "M256F";
      M256A_IDB : Array[0.."CONST_dNumberOfHeadsCycle"] of "M256A";
      M256A_ST_xAllHeadStoppingFaults : Bool;   // Cumulative Head in alarm
      M256F_ST_xAllHeadStoppingFaults : Bool;   // Cumulative Head in alarm
      M256M_ST_xAllHeadStoppingFaults : Bool;   // Cumulative Head in alarm
      M256M_ST_xAllHeadInitialized : Bool;
      M256M_ST_xAllHeadReferred : Bool;
      M256M_ST_xAllHeadPositioned : Bool;
      M256M_ST_xAllHeadIPLinked : Bool;
   END_VAR
   VAR_TEMP
      TMP_rgxHeadReferredSwitch : Array[0.."CONST_dNumberOfHeadsCycle"] of Bool;
      TMP_rgxHeadVirtualCollision : Array[0.."CONST_dNumberOfHeadsCycle"] of Bool;
      TMP_OS_XBrakeRelease : Bool;
      TMP_OS_XBrakeEngage : Bool;
      TMP_xHeadReferredSwicth : Bool;
      TMP_dIndex : DInt;
      TMP_dIndex2Nd : DInt;
      TMP_xDummy : Bool;
   END_VAR
BEGIN

REGION Network 1: #### COSTANTS ####
END_REGION

REGION Network 2: #### ALARMS ####
END_REGION

REGION Network 3: Op. side head overstroke
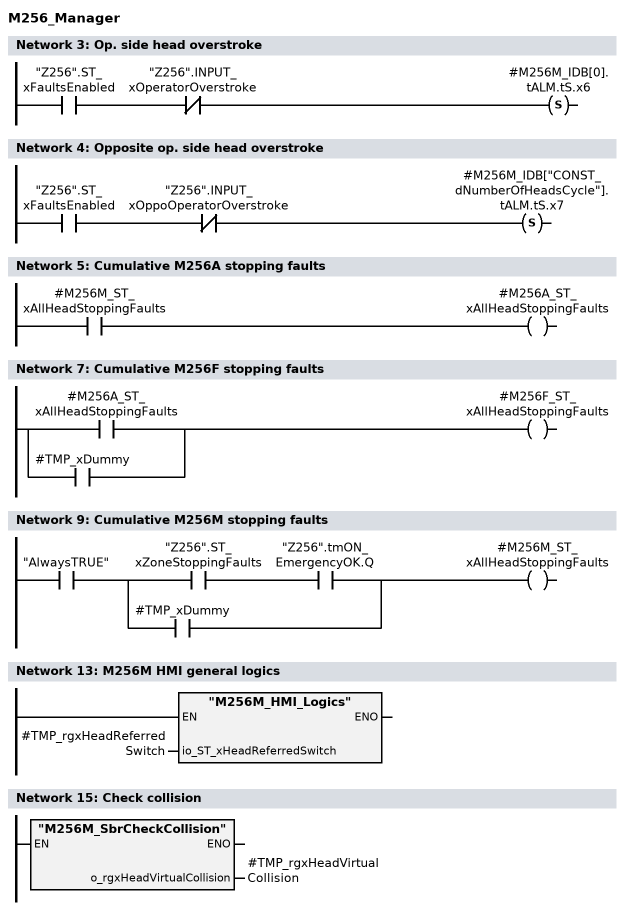
   RUNG wire#powerrail
      Contact( "Z256".ST_xFaultsEnabled )
      I_Contact( "Z256".INPUT_xOperatorOverstroke )
      S_Coil( #M256M_IDB[0].tALM.tS.x6 )
   END_RUNG
   // the same network as SCL:
   IF "Z256".ST_xFaultsEnabled AND NOT "Z256".INPUT_xOperatorOverstroke THEN
       #M256M_IDB[0].tALM.tS.x6 := TRUE;
   END_IF;
END_REGION

REGION Network 4: Opposite op. side head overstroke
   RUNG wire#powerrail
      Contact( "Z256".ST_xFaultsEnabled )
      I_Contact( "Z256".INPUT_xOppoOperatorOverstroke )
      S_Coil( #M256M_IDB["CONST_dNumberOfHeadsCycle"].tALM.tS.x7 )
   END_RUNG
   // the same network as SCL:
   IF "Z256".ST_xFaultsEnabled AND NOT "Z256".INPUT_xOppoOperatorOverstroke THEN
       #M256M_IDB["CONST_dNumberOfHeadsCycle"].tALM.tS.x7 := TRUE;
   END_IF;
END_REGION

REGION Network 5: Cumulative M256A stopping faults
   RUNG wire#powerrail
      Contact( #M256M_ST_xAllHeadStoppingFaults )
      Coil( #M256A_ST_xAllHeadStoppingFaults )
   END_RUNG
   // the same network as SCL:
   #M256A_ST_xAllHeadStoppingFaults := #M256M_ST_xAllHeadStoppingFaults;
END_REGION

REGION Network 6 (SCL): Cumulative M256F faults status
   #TMP_xDummy := FALSE;
   FOR #TMP_dIndex := 0 TO "CONST_dNumberOfHeadsCycle" DO
       IF #M256F_IDB[#TMP_dIndex].ST_xStoppingFaults THEN
           #TMP_xDummy := TRUE;
       END_IF;
   END_FOR;
END_REGION

REGION Network 7: Cumulative M256F stopping faults
   RUNG wire#powerrail
      Contact( #M256A_ST_xAllHeadStoppingFaults )
      wire#w1
      Coil( #M256F_ST_xAllHeadStoppingFaults )
   END_RUNG
   RUNG wire#powerrail
      Contact( #TMP_xDummy )
   END_RUNG wire#w1
   // the same network as SCL:
   #M256F_ST_xAllHeadStoppingFaults := #M256A_ST_xAllHeadStoppingFaults OR #TMP_xDummy;
END_REGION

